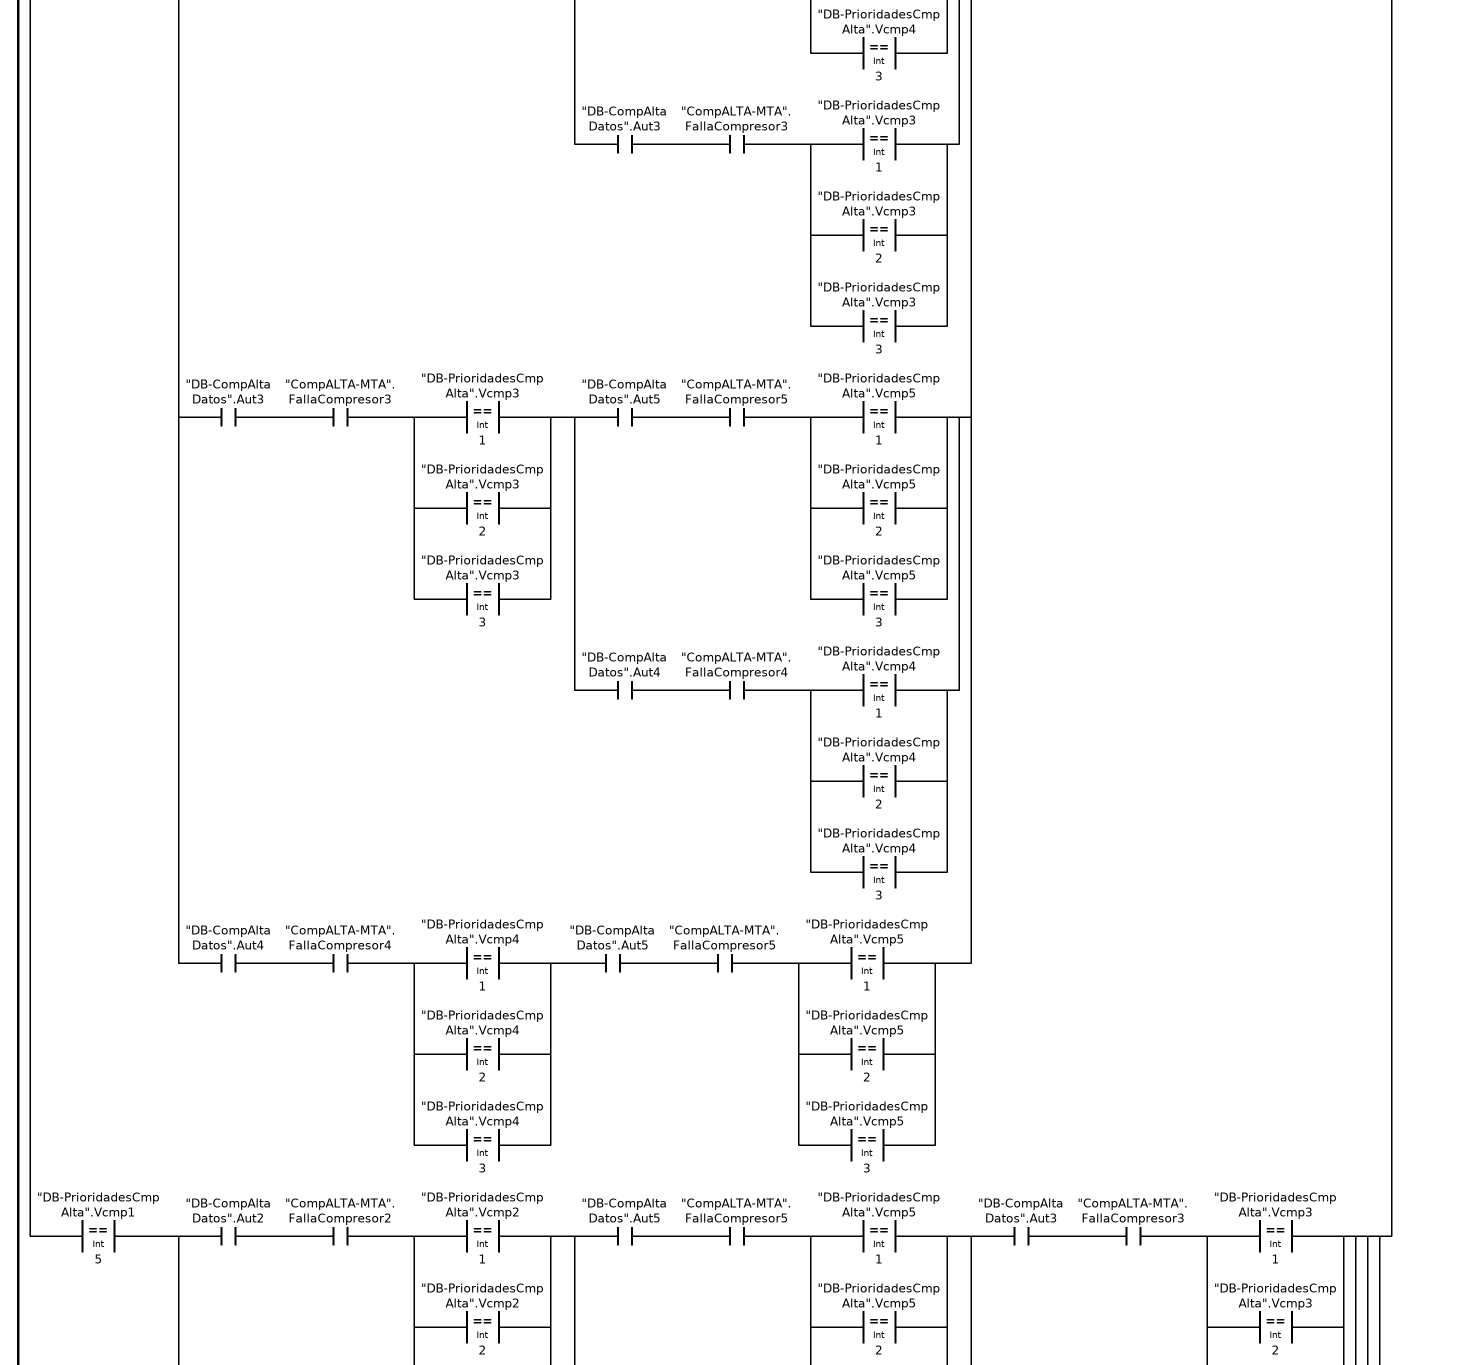
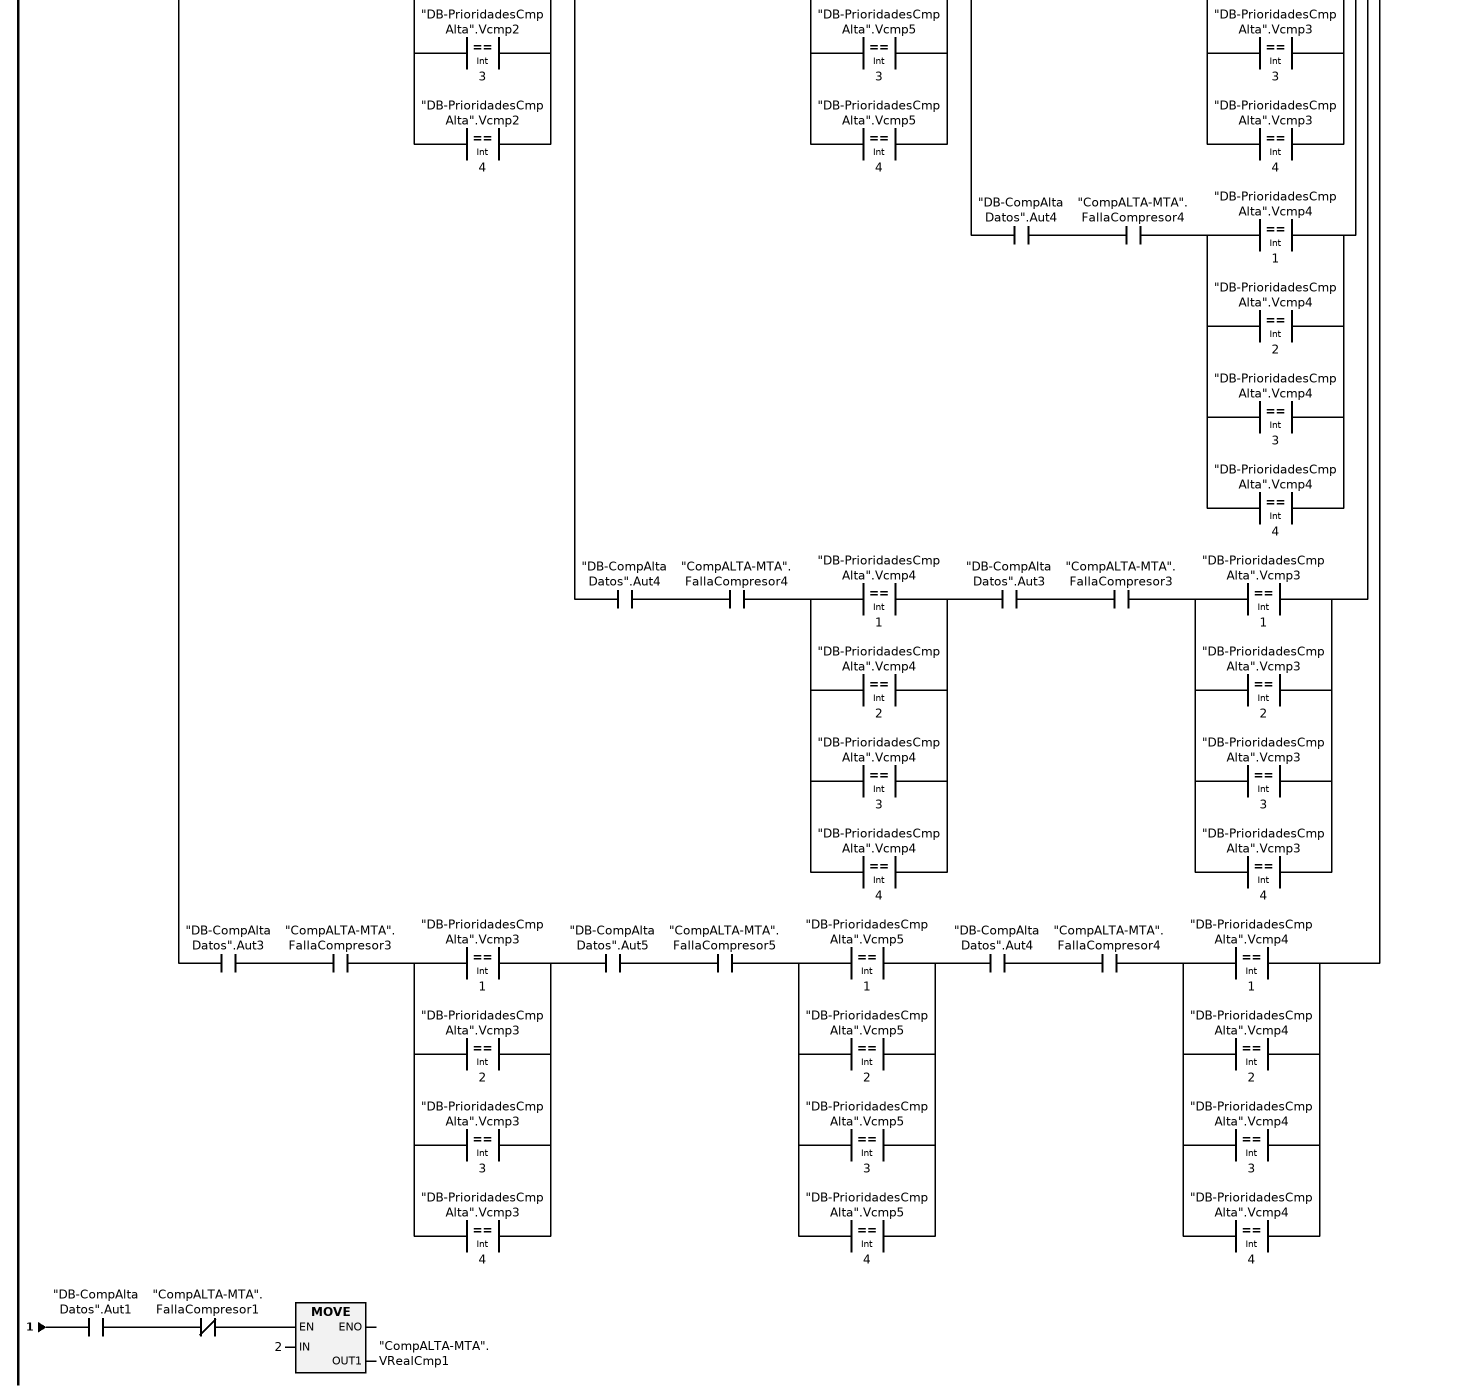
   IF (("DB-PrioridadesCmpAlta".Vcmp1 = 2) OR (("DB-PrioridadesCmpAlta".Vcmp1 = 3) AND (("DB-CompAltaDatos".Aut2 AND "CompALTA-MTA".FallaCompresor2 AND (("DB-PrioridadesCmpAlta".Vcmp2 = 2) OR ("DB-PrioridadesCmpAlta".Vcmp2 = 1))) OR ("DB-CompAltaDatos".Aut3 AND "CompALTA-MTA".FallaCompresor3 AND (("DB-PrioridadesCmpAlta".Vcmp3 = 2) OR ("DB-PrioridadesCmpAlta".Vcmp3 = 1))) OR ("DB-CompAltaDatos".Aut4 AND "CompALTA-MTA".FallaCompresor4 AND (("DB-PrioridadesCmpAlta".Vcmp4 = 2) OR ("DB-PrioridadesCmpAlta".Vcmp4 = 1))) OR ("DB-CompAltaDatos".Aut5 AND "CompALTA-MTA".FallaCompresor5 AND (("DB-PrioridadesCmpAlta".Vcmp5 = 2) OR ("DB-PrioridadesCmpAlta".Vcmp5 = 1))))) OR (("DB-PrioridadesCmpAlta".Vcmp1 = 4) AND (("DB-CompAltaDatos".Aut2 AND "CompALTA-MTA".FallaCompresor2 AND (("DB-PrioridadesCmpAlta".Vcmp2 = 1) OR ("DB-PrioridadesCmpAlta".Vcmp2 = 2) OR ("DB-PrioridadesCmpAlta".Vcmp2 = 3)) AND (("DB-CompAltaDatos".Aut5 AND "CompALTA-MTA".FallaCompresor5 AND (("DB-PrioridadesCmpAlta".Vcmp5 = 1) OR ("DB-PrioridadesCmpAlta".Vcmp5 = 2) OR ("DB-PrioridadesCmpAlta".Vcmp5 = 3))) OR ("DB-CompAltaDatos".Aut4 AND "CompALTA-MTA".FallaCompresor4 AND (("DB-PrioridadesCmpAlta".Vcmp4 = 1) OR ("DB-PrioridadesCmpAlta".Vcmp4 = 2) OR ("DB-PrioridadesCmpAlta".Vcmp4 = 3))) OR ("DB-CompAltaDatos".Aut3 AND "CompALTA-MTA".FallaCompresor3 AND (("DB-PrioridadesCmpAlta".Vcmp3 = 1) OR ("DB-PrioridadesCmpAlta".Vcmp3 = 2) OR ("DB-PrioridadesCmpAlta".Vcmp3 = 3))))) OR ("DB-CompAltaDatos".Aut3 AND "CompALTA-MTA".FallaCompresor3 AND (("DB-PrioridadesCmpAlta".Vcmp3 = 1) OR ("DB-PrioridadesCmpAlta".Vcmp3 = 2) OR ("DB-PrioridadesCmpAlta".Vcmp3 = 3)) AND (("DB-CompAltaDatos".Aut5 AND "CompALTA-MTA".FallaCompresor5 AND (("DB-PrioridadesCmpAlta".Vcmp5 = 1) OR ("DB-PrioridadesCmpAlta".Vcmp5 = 2) OR ("DB-PrioridadesCmpAlta".Vcmp5 = 3))) OR ("DB-CompAltaDatos".Aut4 AND "CompALTA-MTA".FallaCompresor4 AND (("DB-PrioridadesCmpAlta".Vcmp4 = 1) OR ("DB-PrioridadesCmpAlta".Vcmp4 = 2) OR ("DB-PrioridadesCmpAlta".Vcmp4 = 3))))) OR ("DB-CompAltaDatos".Aut4 AND "CompALTA-MTA".FallaCompresor4 AND (("DB-PrioridadesCmpAlta".Vcmp4 = 1) OR ("DB-PrioridadesCmpAlta".Vcmp4 = 2) OR ("DB-PrioridadesCmpAlta".Vcmp4 = 3)) AND "DB-CompAltaDatos".Aut5 AND "CompALTA-MTA".FallaCompresor5 AND (("DB-PrioridadesCmpAlta".Vcmp5 = 1) OR ("DB-PrioridadesCmpAlta".Vcmp5 = 2) OR ("DB-PrioridadesCmpAlta".Vcmp5 = 3))))) OR (("DB-PrioridadesCmpAlta".Vcmp1 = 5) AND (("DB-CompAltaDatos".Aut2 AND "CompALTA-MTA".FallaCompresor2 AND (("DB-PrioridadesCmpAlta".Vcmp2 = 1) OR ("DB-PrioridadesCmpAlta".Vcmp2 = 2) OR ("DB-PrioridadesCmpAlta".Vcmp2 = 3) OR ("DB-PrioridadesCmpAlta".Vcmp2 = 4)) AND (("DB-CompAltaDatos".Aut5 AND "CompALTA-MTA".FallaCompresor5 AND (("DB-PrioridadesCmpAlta".Vcmp5 = 1) OR ("DB-PrioridadesCmpAlta".Vcmp5 = 2) OR ("DB-PrioridadesCmpAlta".Vcmp5 = 3) OR ("DB-PrioridadesCmpAlta".Vcmp5 = 4)) AND (("DB-CompAltaDatos".Aut3 AND "CompALTA-MTA".FallaCompresor3 AND (("DB-PrioridadesCmpAlta".Vcmp3 = 1) OR ("DB-PrioridadesCmpAlta".Vcmp3 = 2) OR ("DB-PrioridadesCmpAlta".Vcmp3 = 3) OR ("DB-PrioridadesCmpAlta".Vcmp3 = 4))) OR ("DB-CompAltaDatos".Aut4 AND "CompALTA-MTA".FallaCompresor4 AND (("DB-PrioridadesCmpAlta".Vcmp4 = 1) OR ("DB-PrioridadesCmpAlta".Vcmp4 = 2) OR ("DB-PrioridadesCmpAlta".Vcmp4 = 3) OR ("DB-PrioridadesCmpAlta".Vcmp4 = 4))))) OR ("DB-CompAltaDatos".Aut4 AND "CompALTA-MTA".FallaCompresor4 AND (("DB-PrioridadesCmpAlta".Vcmp4 = 1) OR ("DB-PrioridadesCmpAlta".Vcmp4 = 2) OR ("DB-PrioridadesCmpAlta".Vcmp4 = 3) OR ("DB-PrioridadesCmpAlta".Vcmp4 = 4)) AND "DB-CompAltaDatos".Aut3 AND "CompALTA-MTA".FallaCompresor3 AND (("DB-PrioridadesCmpAlta".Vcmp3 = 1) OR ("DB-PrioridadesCmpAlta".Vcmp3 = 2) OR ("DB-PrioridadesCmpAlta".Vcmp3 = 3) OR ("DB-PrioridadesCmpAlta".Vcmp3 = 4))))) OR ("DB-CompAltaDatos".Aut3 AND "CompALTA-MTA".FallaCompresor3 AND (("DB-PrioridadesCmpAlta".Vcmp3 = 1) OR ("DB-PrioridadesCmpAlta".Vcmp3 = 2) OR ("DB-PrioridadesCmpAlta".Vcmp3 = 3) OR ("DB-PrioridadesCmpAlta".Vcmp3 = 4)) AND "DB-CompAltaDatos".Aut5 AND "CompALTA-MTA".FallaCompresor5 AND (("DB-PrioridadesCmpAlta".Vcmp5 = 1) OR ("DB-PrioridadesCmpAlta".Vcmp5 = 2) OR ("DB-PrioridadesCmpAlta".Vcmp5 = 3) OR ("DB-PrioridadesCmpAlta".Vcmp5 = 4)) AND "DB-CompAltaDatos".Aut4 AND "CompALTA-MTA".FallaCompresor4 AND (("DB-PrioridadesCmpAlta".Vcmp4 = 1) OR ("DB-PrioridadesCmpAlta".Vcmp4 = 2) OR ("DB-PrioridadesCmpAlta".Vcmp4 = 3) OR ("DB-PrioridadesCmpAlta".Vcmp4 = 4)))))) AND "DB-CompAltaDatos".Aut1 AND NOT "CompALTA-MTA".FallaCompresor1 THEN
       "CompALTA-MTA".VRealCmp1 := 2;
   END_IF;
END_REGION

REGION Network 5
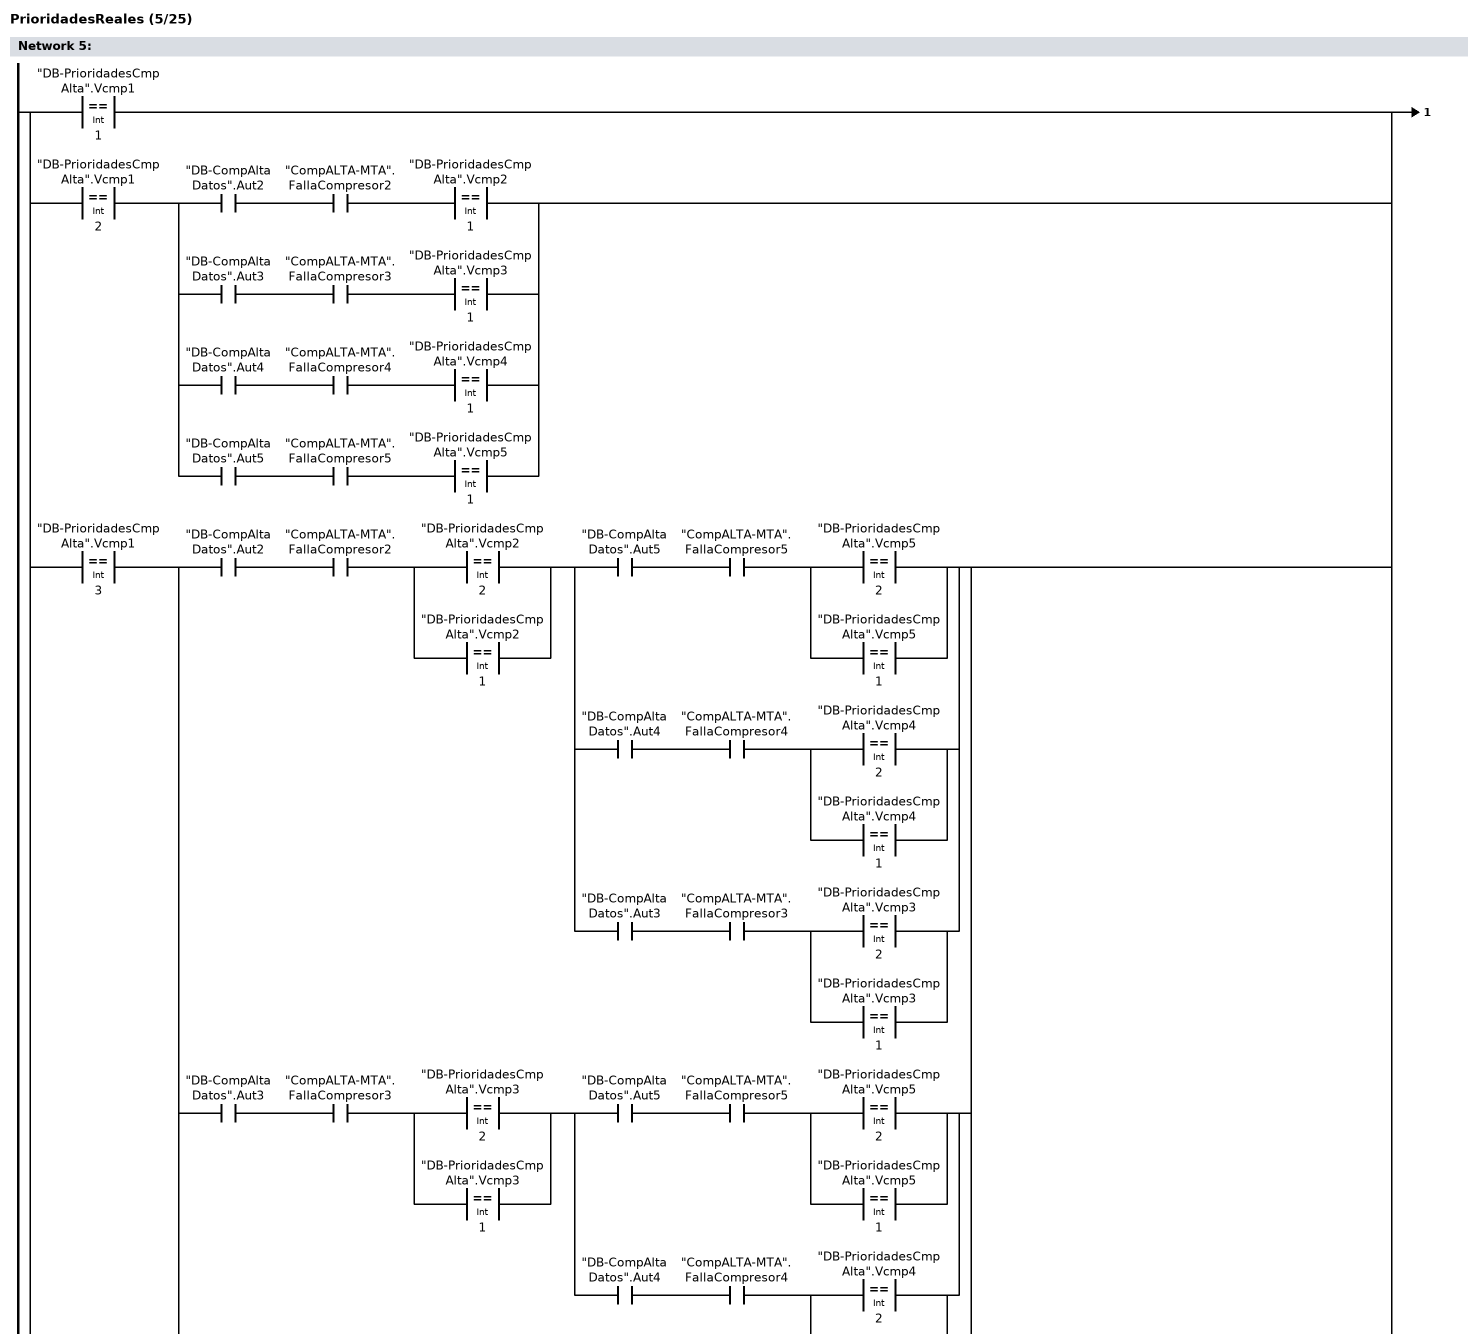
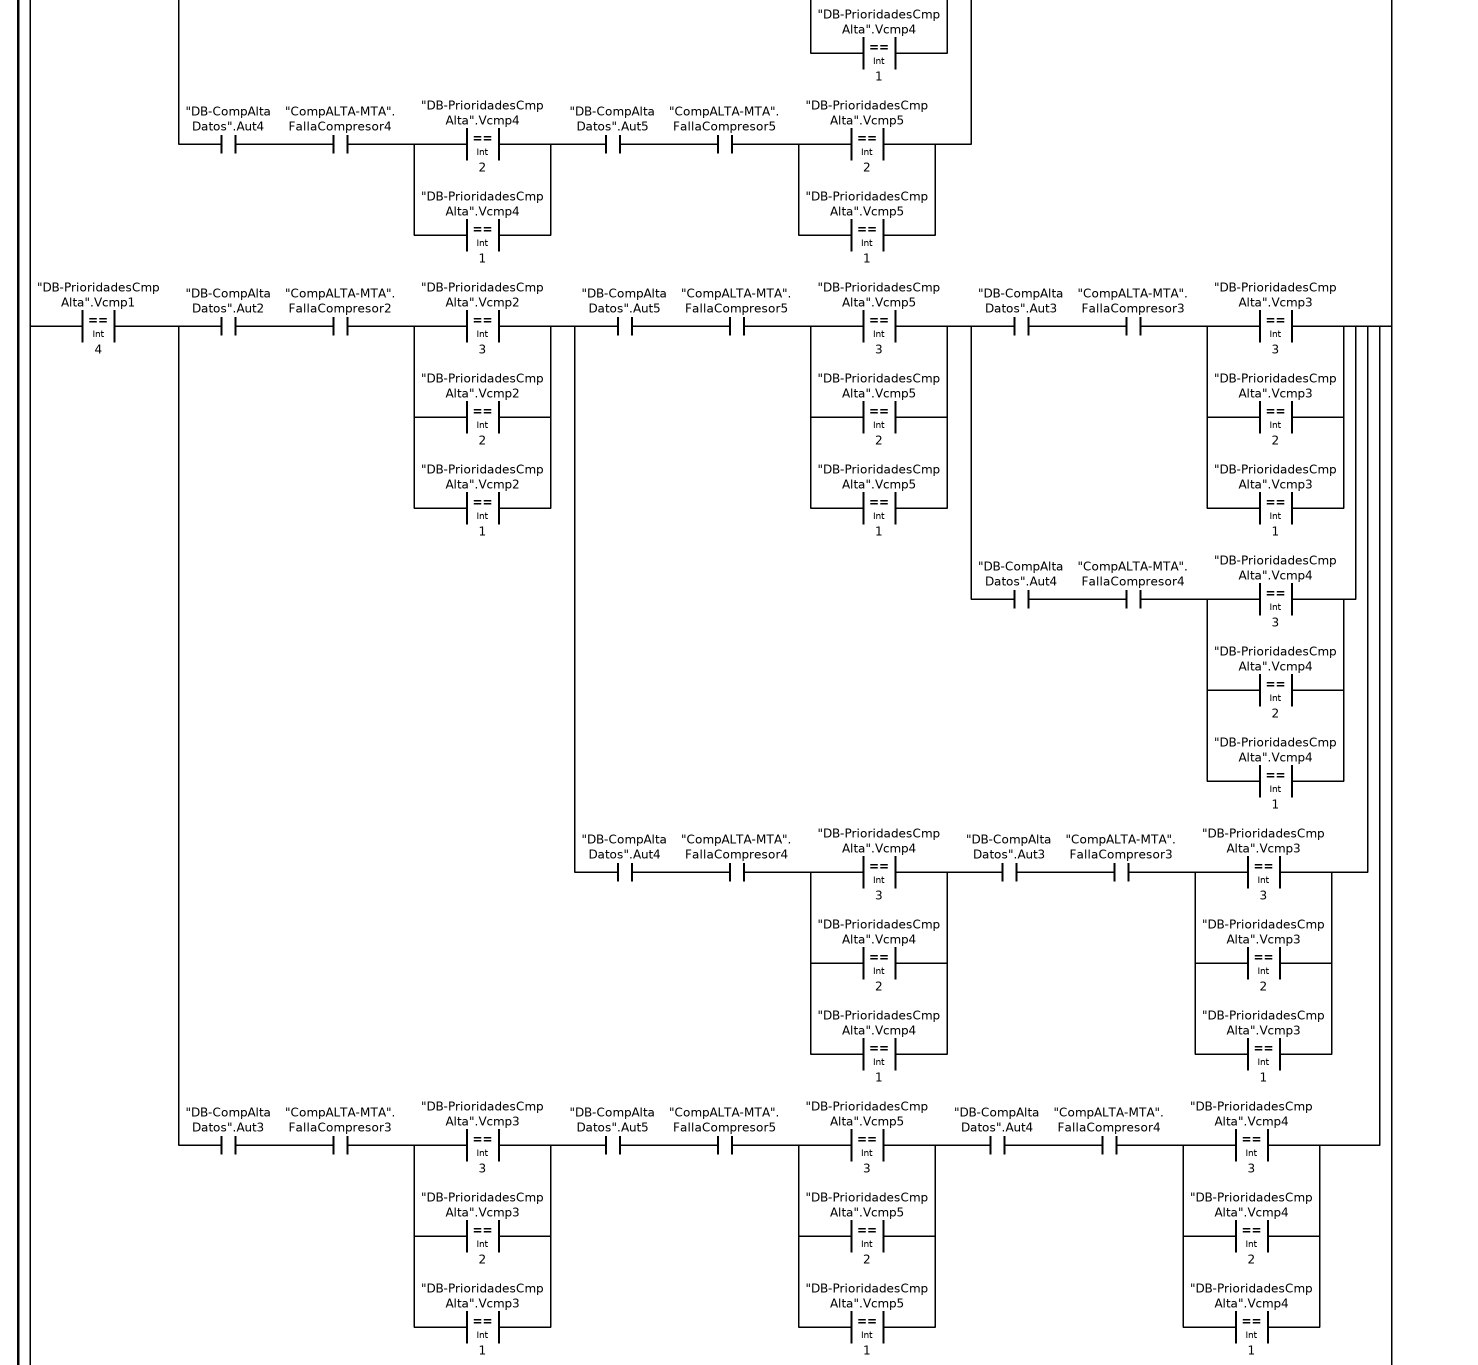
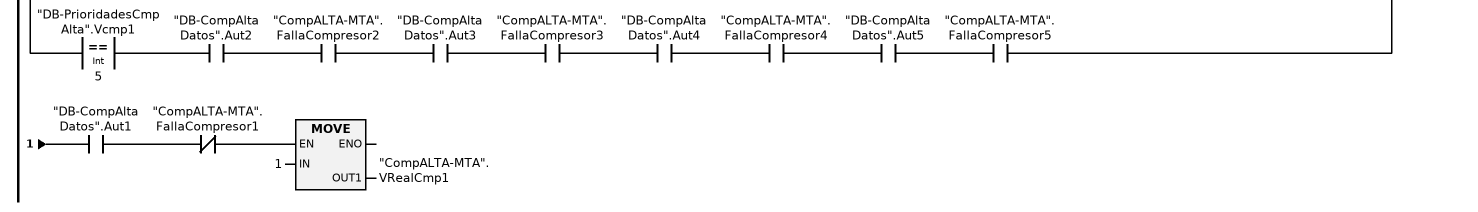
   IF (("DB-PrioridadesCmpAlta".Vcmp1 = 1) OR (("DB-PrioridadesCmpAlta".Vcmp1 = 2) AND (("DB-CompAltaDatos".Aut2 AND "CompALTA-MTA".FallaCompresor2 AND ("DB-PrioridadesCmpAlta".Vcmp2 = 1)) OR ("DB-CompAltaDatos".Aut3 AND "CompALTA-MTA".FallaCompresor3 AND ("DB-PrioridadesCmpAlta".Vcmp3 = 1)) OR ("DB-CompAltaDatos".Aut4 AND "CompALTA-MTA".FallaCompresor4 AND ("DB-PrioridadesCmpAlta".Vcmp4 = 1)) OR ("DB-CompAltaDatos".Aut5 AND "CompALTA-MTA".FallaCompresor5 AND ("DB-PrioridadesCmpAlta".Vcmp5 = 1)))) OR (("DB-PrioridadesCmpAlta".Vcmp1 = 3) AND (("DB-CompAltaDatos".Aut2 AND "CompALTA-MTA".FallaCompresor2 AND (("DB-PrioridadesCmpAlta".Vcmp2 = 2) OR ("DB-PrioridadesCmpAlta".Vcmp2 = 1)) AND (("DB-CompAltaDatos".Aut5 AND "CompALTA-MTA".FallaCompresor5 AND (("DB-PrioridadesCmpAlta".Vcmp5 = 2) OR ("DB-PrioridadesCmpAlta".Vcmp5 = 1))) OR ("DB-CompAltaDatos".Aut4 AND "CompALTA-MTA".FallaCompresor4 AND (("DB-PrioridadesCmpAlta".Vcmp4 = 2) OR ("DB-PrioridadesCmpAlta".Vcmp4 = 1))) OR ("DB-CompAltaDatos".Aut3 AND "CompALTA-MTA".FallaCompresor3 AND (("DB-PrioridadesCmpAlta".Vcmp3 = 2) OR ("DB-PrioridadesCmpAlta".Vcmp3 = 1))))) OR ("DB-CompAltaDatos".Aut3 AND "CompALTA-MTA".FallaCompresor3 AND (("DB-PrioridadesCmpAlta".Vcmp3 = 2) OR ("DB-PrioridadesCmpAlta".Vcmp3 = 1)) AND (("DB-CompAltaDatos".Aut5 AND "CompALTA-MTA".FallaCompresor5 AND (("DB-PrioridadesCmpAlta".Vcmp5 = 2) OR ("DB-PrioridadesCmpAlta".Vcmp5 = 1))) OR ("DB-CompAltaDatos".Aut4 AND "CompALTA-MTA".FallaCompresor4 AND (("DB-PrioridadesCmpAlta".Vcmp4 = 2) OR ("DB-PrioridadesCmpAlta".Vcmp4 = 1))))) OR ("DB-CompAltaDatos".Aut4 AND "CompALTA-MTA".FallaCompresor4 AND (("DB-PrioridadesCmpAlta".Vcmp4 = 2) OR ("DB-PrioridadesCmpAlta".Vcmp4 = 1)) AND "DB-CompAltaDatos".Aut5 AND "CompALTA-MTA".FallaCompresor5 AND (("DB-PrioridadesCmpAlta".Vcmp5 = 2) OR ("DB-PrioridadesCmpAlta".Vcmp5 = 1))))) OR (("DB-PrioridadesCmpAlta".Vcmp1 = 4) AND (("DB-CompAltaDatos".Aut2 AND "CompALTA-MTA".FallaCompresor2 AND (("DB-PrioridadesCmpAlta".Vcmp2 = 3) OR ("DB-PrioridadesCmpAlta".Vcmp2 = 2) OR ("DB-PrioridadesCmpAlta".Vcmp2 = 1)) AND (("DB-CompAltaDatos".Aut5 AND "CompALTA-MTA".FallaCompresor5 AND (("DB-PrioridadesCmpAlta".Vcmp5 = 3) OR ("DB-PrioridadesCmpAlta".Vcmp5 = 2) OR ("DB-PrioridadesCmpAlta".Vcmp5 = 1)) AND (("DB-CompAltaDatos".Aut3 AND "CompALTA-MTA".FallaCompresor3 AND (("DB-PrioridadesCmpAlta".Vcmp3 = 3) OR ("DB-PrioridadesCmpAlta".Vcmp3 = 2) OR ("DB-PrioridadesCmpAlta".Vcmp3 = 1))) OR ("DB-CompAltaDatos".Aut4 AND "CompALTA-MTA".FallaCompresor4 AND (("DB-PrioridadesCmpAlta".Vcmp4 = 3) OR ("DB-PrioridadesCmpAlta".Vcmp4 = 2) OR ("DB-PrioridadesCmpAlta".Vcmp4 = 1))))) OR ("DB-CompAltaDatos".Aut4 AND "CompALTA-MTA".FallaCompresor4 AND (("DB-PrioridadesCmpAlta".Vcmp4 = 3) OR ("DB-PrioridadesCmpAlta".Vcmp4 = 2) OR ("DB-PrioridadesCmpAlta".Vcmp4 = 1)) AND "DB-CompAltaDatos".Aut3 AND "CompALTA-MTA".FallaCompresor3 AND (("DB-PrioridadesCmpAlta".Vcmp3 = 3) OR ("DB-PrioridadesCmpAlta".Vcmp3 = 2) OR ("DB-PrioridadesCmpAlta".Vcmp3 = 1))))) OR ("DB-CompAltaDatos".Aut3 AND "CompALTA-MTA".FallaCompresor3 AND (("DB-PrioridadesCmpAlta".Vcmp3 = 3) OR ("DB-PrioridadesCmpAlta".Vcmp3 = 2) OR ("DB-PrioridadesCmpAlta".Vcmp3 = 1)) AND "DB-CompAltaDatos".Aut5 AND "CompALTA-MTA".FallaCompresor5 AND (("DB-PrioridadesCmpAlta".Vcmp5 = 3) OR ("DB-PrioridadesCmpAlta".Vcmp5 = 2) OR ("DB-PrioridadesCmpAlta".Vcmp5 = 1)) AND "DB-CompAltaDatos".Aut4 AND "CompALTA-MTA".FallaCompresor4 AND (("DB-PrioridadesCmpAlta".Vcmp4 = 3) OR ("DB-PrioridadesCmpAlta".Vcmp4 = 2) OR ("DB-PrioridadesCmpAlta".Vcmp4 = 1))))) OR (("DB-PrioridadesCmpAlta".Vcmp1 = 5) AND "DB-CompAltaDatos".Aut2 AND "CompALTA-MTA".FallaCompresor2 AND "DB-CompAltaDatos".Aut3 AND "CompALTA-MTA".FallaCompresor3 AND "DB-CompAltaDatos".Aut4 AND "CompALTA-MTA".FallaCompresor4 AND "DB-CompAltaDatos".Aut5 AND "CompALTA-MTA".FallaCompresor5)) AND "DB-CompAltaDatos".Aut1 AND NOT "CompALTA-MTA".FallaCompresor1 THEN
       "CompALTA-MTA".VRealCmp1 := 1;
   END_IF;
END_REGION

REGION Network 8
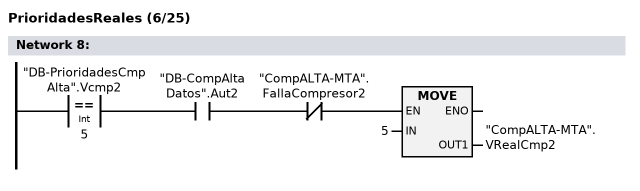
   RUNG wire#powerrail
      { S7_Templates := "SrcType := Int" } EQ_Contact(in1 := "DB-PrioridadesCmpAlta".Vcmp2, in2 := 5)
      Contact( "DB-CompAltaDatos".Aut2 )
      I_Contact( "CompALTA-MTA".FallaCompresor2 )
      { S7_GenerateENO := "TRUE" } Move(in := 5, out1 => "CompALTA-MTA".VRealCmp2)
   END_RUNG
   // the same network as SCL:
   IF ("DB-PrioridadesCmpAlta".Vcmp2 = 5) AND "DB-CompAltaDatos".Aut2 AND NOT "CompALTA-MTA".FallaCompresor2 THEN
       "CompALTA-MTA".VRealCmp2 := 5;
   END_IF;
END_REGION

REGION Network 9
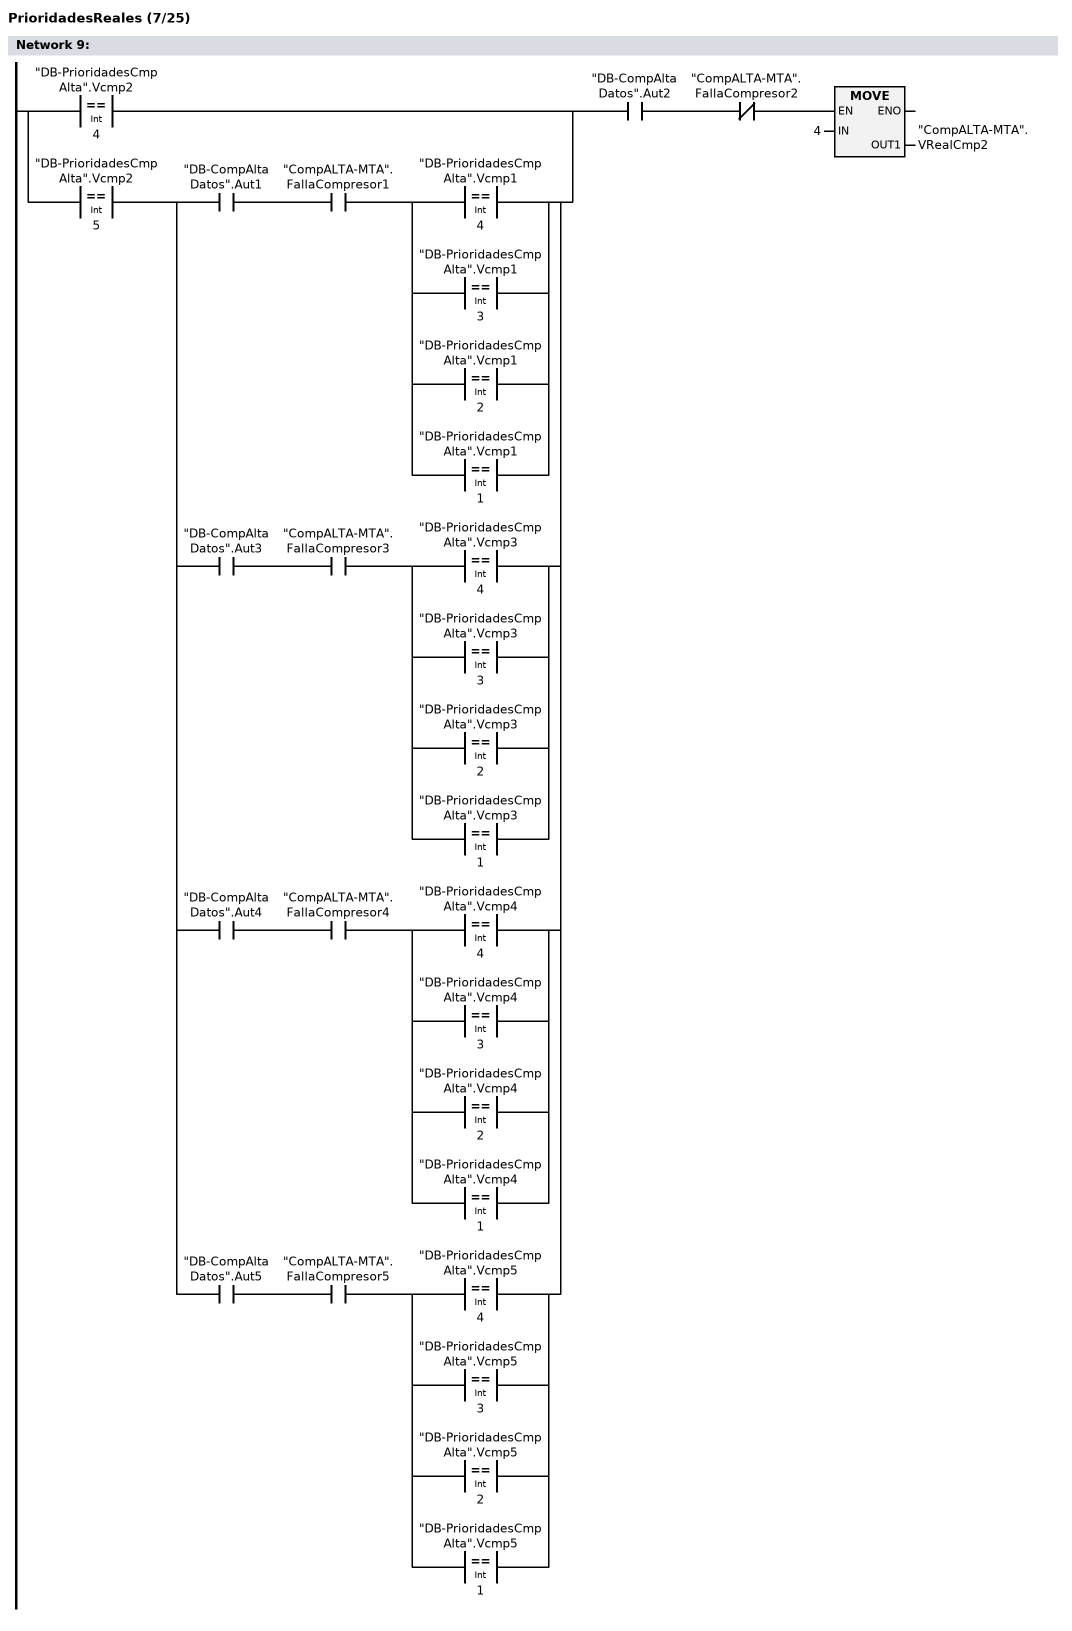
   IF (("DB-PrioridadesCmpAlta".Vcmp2 = 4) OR (("DB-PrioridadesCmpAlta".Vcmp2 = 5) AND (("DB-CompAltaDatos".Aut1 AND "CompALTA-MTA".FallaCompresor1 AND (("DB-PrioridadesCmpAlta".Vcmp1 = 4) OR ("DB-PrioridadesCmpAlta".Vcmp1 = 3) OR ("DB-PrioridadesCmpAlta".Vcmp1 = 2) OR ("DB-PrioridadesCmpAlta".Vcmp1 = 1))) OR ("DB-CompAltaDatos".Aut3 AND "CompALTA-MTA".FallaCompresor3 AND (("DB-PrioridadesCmpAlta".Vcmp3 = 4) OR ("DB-PrioridadesCmpAlta".Vcmp3 = 3) OR ("DB-PrioridadesCmpAlta".Vcmp3 = 2) OR ("DB-PrioridadesCmpAlta".Vcmp3 = 1))) OR ("DB-CompAltaDatos".Aut4 AND "CompALTA-MTA".FallaCompresor4 AND (("DB-PrioridadesCmpAlta".Vcmp4 = 4) OR ("DB-PrioridadesCmpAlta".Vcmp4 = 3) OR ("DB-PrioridadesCmpAlta".Vcmp4 = 2) OR ("DB-PrioridadesCmpAlta".Vcmp4 = 1))) OR ("DB-CompAltaDatos".Aut5 AND "CompALTA-MTA".FallaCompresor5 AND (("DB-PrioridadesCmpAlta".Vcmp5 = 4) OR ("DB-PrioridadesCmpAlta".Vcmp5 = 3) OR ("DB-PrioridadesCmpAlta".Vcmp5 = 2) OR ("DB-PrioridadesCmpAlta".Vcmp5 = 1)))))) AND "DB-CompAltaDatos".Aut2 AND NOT "CompALTA-MTA".FallaCompresor2 THEN
       "CompALTA-MTA".VRealCmp2 := 4;
   END_IF;
END_REGION

REGION Network 10
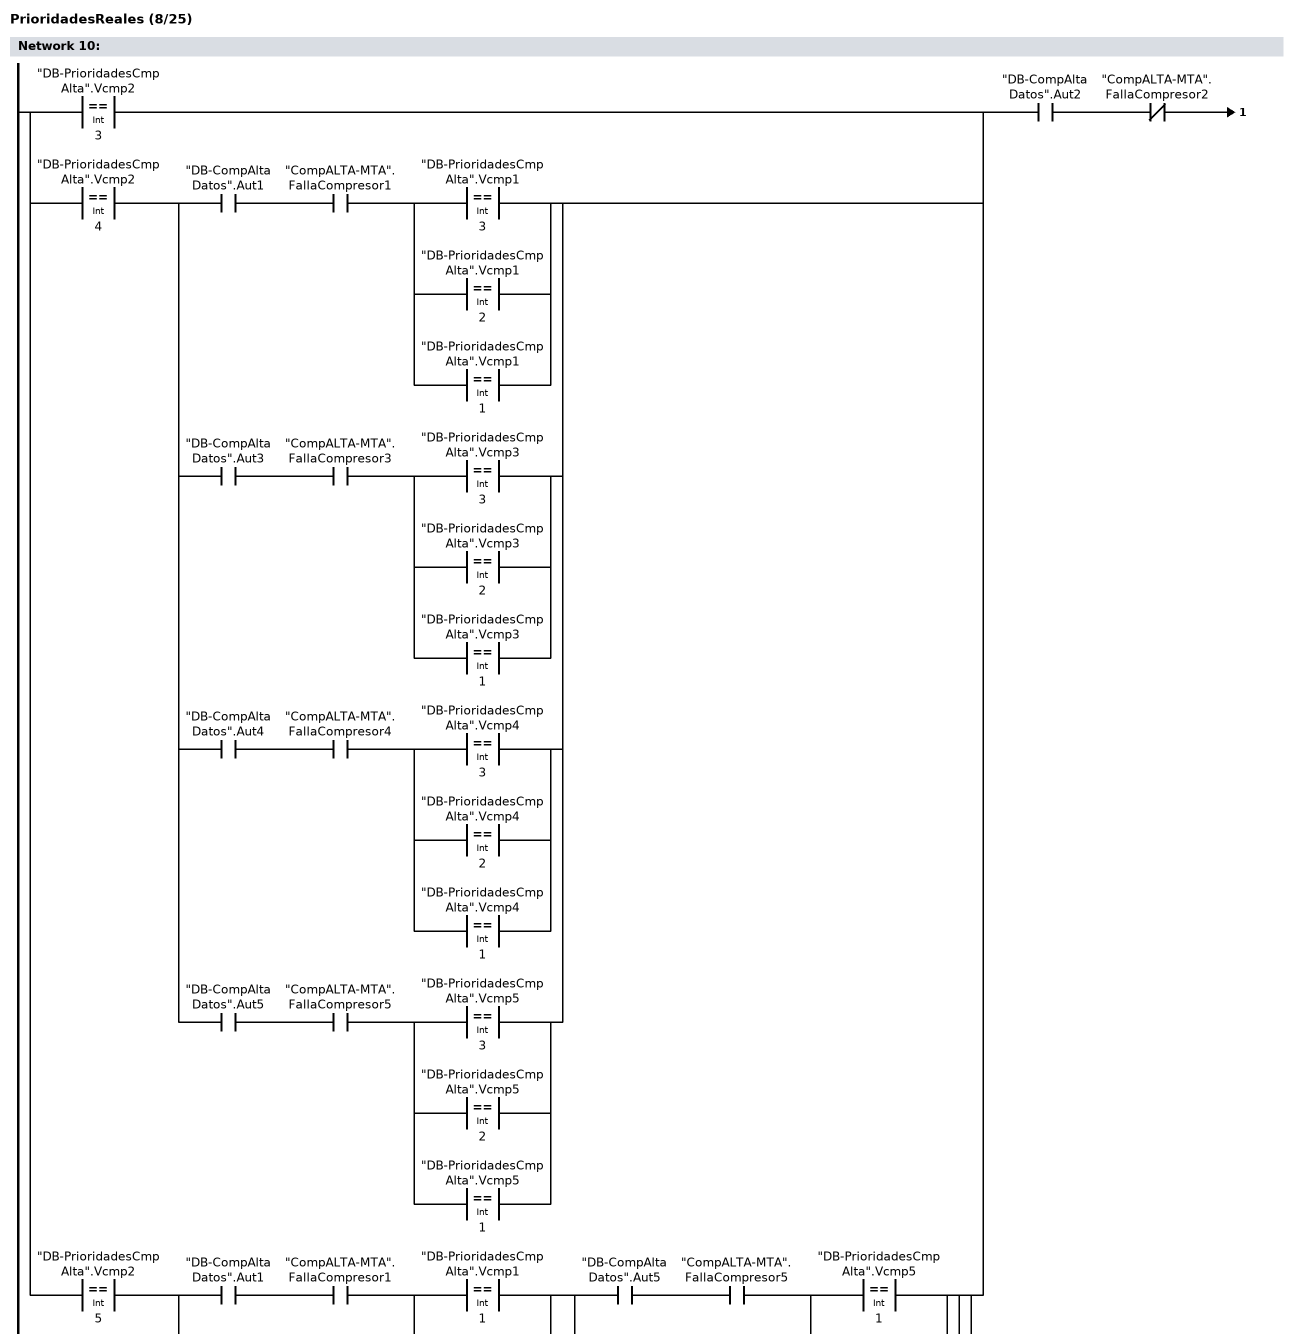
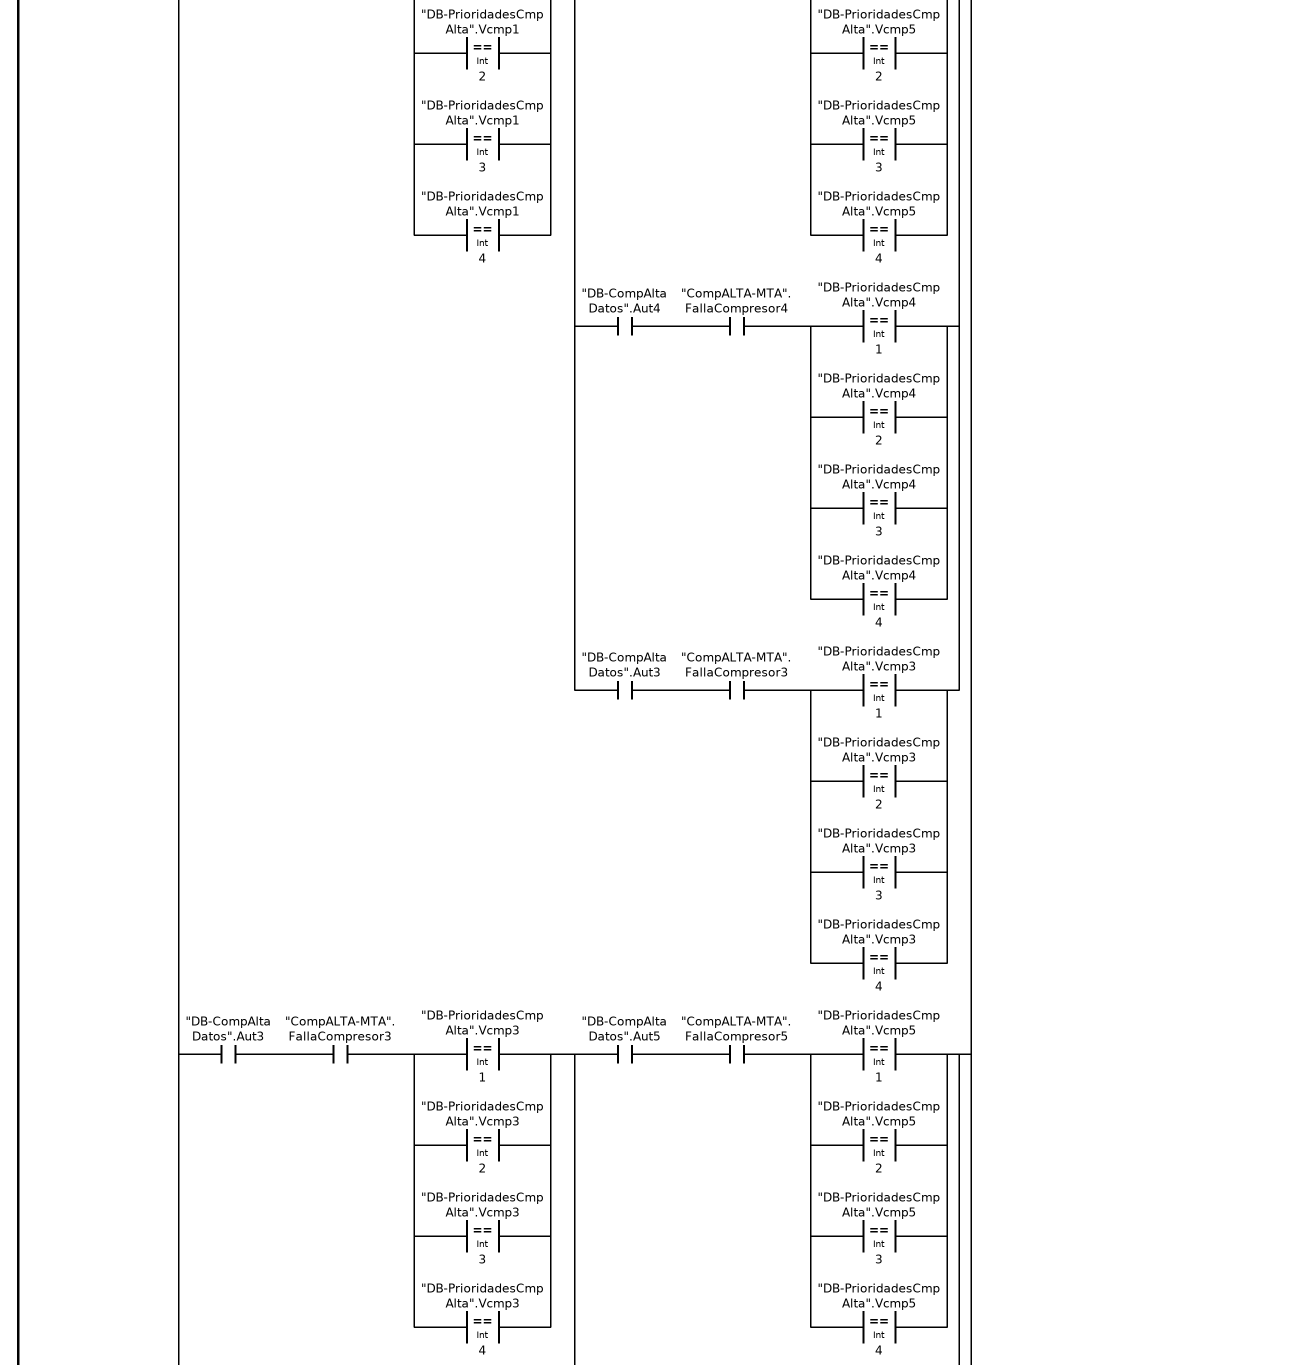
